HMI tags "Tabla de variables estándar"
   "IndR6" : Bool AT %DB121.DBX3.0, 100 ms
   "IndVparp6" : Bool AT %DB121.DBX70.5, 1 s
   "Auto6" : Bool AT %DB88.DBX10.5, 1 s
   "PanMCH6" : Bool AT %DB88.DBX6.5, 1 s
   "LimSUP6" : Real AT %DB122.DBD20, 1 s
   "LimINF6" : Real AT %DB122.DBD44, 1 s
   "VCMP6" : Int AT %DB125.DBW12, 1 s
   "IncP6" : Bool AT %DB125.DBX16.1, 100 ms
   "DecP6" : Bool AT %DB125.DBX16.7, 1 s
   "SPONF6" : Real AT %DB136.DBD24, 1 s
   "SPOFFF6" : Real AT %DB136.DBD48, 1 s
   "ForzarMarcha6" : Bool AT %DB136.DBX0.5, 1 s
   "ForzarParada6" : Bool AT %DB136.DBX1.3, 1 s
   "ForzandoMarcha6" : Bool AT %DB136.DBX2.1, 1 s
   "SPON6" : Real AT %DB135.DBD32, 1 s
   "SPOFF6" : Real AT %DB135.DBD56, 1 s
   "AnimMenuMC006" : Int AT %DB135.DBW10, 1 s
   "MantMC006" : Bool AT %DB135.DBX60.5, 1 s
   "MarchaOK6" : Bool AT %DB135.DBX61.3, 1 s
   "MarchaMC006" : Bool AT %DB135.DBX62.1, 1 s
   "ParadaMC006" : Bool AT %DB135.DBX62.7, 1 s
   "HORAS6" : DInt AT %DB73.DBD20, 1 s
   "MIN6" : Int AT %DB73.DBW34, 1 s
   "AnimMotorMC006" : Byte AT %DB46.DBB45, 1 s
   "EV6" : Bool AT %Q6.3, 1 s
   "ProxMantMC001_1" : DInt = PLC ProxMantMC001_1 AT %MD768, 1 s
   "ProxMantMC001_2" : DInt = PLC ProxMantMC001_2 AT %MD792, 1 s
   "Varios_UltimoMantMC001_1" : DInt = PLC Varios.UltimoMantMC001_1 AT %DB2.DBD48, 1 s
   "Varios_UltimoMantMC001_2" : DInt = PLC Varios.UltimoMantMC001_2 AT %DB2.DBD72, 1 s
   "ProxMantMC002_1" : DInt = PLC ProxMantMC002_1 AT %MD772, 1 s
   "ProxMantMC002_2" : DInt = PLC ProxMantMC002_2 AT %MD796, 1 s
   "ProxMantMC003_1" : DInt = PLC ProxMantMC003_1 AT %MD776, 1 s
   "ProxMantMC003_2" : DInt = PLC ProxMantMC003_2 AT %MD800, 1 s
   "ProxMantMC004_1" : DInt = PLC ProxMantMC004_1 AT %MD780, 1 s
   "ProxMantMC004_2" : DInt = PLC ProxMantMC004_2 AT %MD804, 1 s
   "ProxMantMC005_1" : DInt = PLC ProxMantMC005_1 AT %MD784, 1 s
   "ProxMantMC005_2" : DInt = PLC ProxMantMC005_2 AT %MD808, 1 s
   "ProxMantMC006_1" : DInt = PLC ProxMantMC006_1 AT %MD788, 1 s
   "ProxMantMC006_2" : DInt = PLC ProxMantMC006_2 AT %MD812, 1 s
   "Varios_UltimoMantMC002_1" : DInt = PLC Varios.UltimoMantMC002_1 AT %DB2.DBD52, 1 s
   "Varios_UltimoMantMC002_2" : DInt = PLC Varios.UltimoMantMC002_2 AT %DB2.DBD76, 1 s
   "Varios_UltimoMantMC003_1" : DInt = PLC Varios.UltimoMantMC003_1 AT %DB2.DBD56, 1 s
   "Varios_UltimoMantMC003_2" : DInt = PLC Varios.UltimoMantMC003_2 AT %DB2.DBD80, 1 s
   "Varios_UltimoMantMC004_1" : DInt = PLC Varios.UltimoMantMC004_1 AT %DB2.DBD60, 1 s
   "Varios_UltimoMantMC004_2" : DInt = PLC Varios.UltimoMantMC004_2 AT %DB2.DBD84, 1 s
   "Varios_UltimoMantMC005_1" : DInt = PLC Varios.UltimoMantMC005_1 AT %DB2.DBD64, 1 s
   "Varios_UltimoMantMC005_2" : DInt = PLC Varios.UltimoMantMC005_2 AT %DB2.DBD88, 1 s
   "Varios_UltimoMantMC006_1" : DInt = PLC Varios.UltimoMantMC006_1 AT %DB2.DBD68, 1 s
   "Varios_UltimoMantMC006_2" : DInt = PLC Varios.UltimoMantMC006_2 AT %DB2.DBD92, 1 s
   "Varios_HorasMantMC001_1" : DInt = PLC Varios.HorasMantMC001_1 AT %DB2.DBD0, 1 s
   "Varios_HorasMantMC006_1" : DInt = PLC Varios.HorasMantMC006_1 AT %DB2.DBD20, 1 s
   "Varios_HorasMantMC006_2" : DInt = PLC Varios.HorasMantMC006_2 AT %DB2.DBD44, 1 s
   "Varios_HorasMantMC002_1" : DInt = PLC Varios.HorasMantMC002_1 AT %DB2.DBD4, 1 s
   "Varios_HorasMantMC001_2" : DInt = PLC Varios.HorasMantMC001_2 AT %DB2.DBD24, 1 s
   "Varios_HorasMantMC002_2" : DInt = PLC Varios.HorasMantMC002_2 AT %DB2.DBD28, 1 s
   "Varios_HorasMantMC004_1" : DInt = PLC Varios.HorasMantMC004_1 AT %DB2.DBD12, 1 s
   "Varios_HorasMantMC004_2" : DInt = PLC Varios.HorasMantMC004_2 AT %DB2.DBD36, 1 s
   "Varios_HorasMantMC005_1" : DInt = PLC Varios.HorasMantMC005_1 AT %DB2.DBD16, 1 s
   "Varios_HorasMantMC005_2" : DInt = PLC Varios.HorasMantMC005_2 AT %DB2.DBD40, 1 s
   "Varios_HorasMantMC003_1" : DInt = PLC Varios.HorasMantMC003_1 AT %DB2.DBD8, 1 s
   "Varios_HorasMantMC003_2" : DInt = PLC Varios.HorasMantMC003_2 AT %DB2.DBD32, 1 s
   "EstadoMantMC003" : Byte = PLC EstadoMantMC003 AT %MB763, 1 s
   "EstadoMantMC005" : Byte = PLC EstadoMantMC005 AT %MB765, 1 s
   "EstadoMantMC004" : Byte = PLC EstadoMantMC004 AT %MB764, 1 s
   "EstadoMantMC002" : Byte = PLC EstadoMantMC002 AT %MB762, 1 s
   "EstadoMantMC001" : Byte = PLC EstadoMantMC001 AT %MB761, 1 s
   "EstadoMantMC006" : Byte = PLC EstadoMantMC006 AT %MB766, 1 s
   "LimiteMantMC001_1" : Bool = PLC LimiteMantMC001_1 AT %M761.0, 1 s
   "LimiteMantMC001_2" : Bool = PLC LimiteMantMC001_2 AT %M761.1, 1 s
   "LimiteMantMC002_1" : Bool = PLC LimiteMantMC002_1 AT %M762.0, 1 s
   "LimiteMantMC002_2" : Bool = PLC LimiteMantMC002_2 AT %M762.1, 1 s
   "LimiteMantMC003_1" : Bool = PLC LimiteMantMC003_1 AT %M763.0, 1 s
   "LimiteMantMC003_2" : Bool = PLC LimiteMantMC003_2 AT %M763.1, 1 s
   "LimiteMantMC004_1" : Bool = PLC LimiteMantMC004_1 AT %M764.0, 1 s
   "LimiteMantMC004_2" : Bool = PLC LimiteMantMC004_2 AT %M764.1, 1 s
   "LimiteMantMC005_1" : Bool = PLC LimiteMantMC005_1 AT %M765.0, 1 s
   "LimiteMantMC005_2" : Bool = PLC LimiteMantMC005_2 AT %M765.1, 1 s
   "LimiteMantMC006_1" : Bool = PLC LimiteMantMC006_1 AT %M766.0, 1 s
   "LimiteMantMC006_2" : Bool = PLC LimiteMantMC006_2 AT %M766.1, 1 s
   "Varios_HorasMantMS050" : DInt = PLC Varios.HorasMantMS050 AT %DB2.DBD96, 1 s
   "Varios_HorasMantMS051" : DInt = PLC Varios.HorasMantMS051 AT %DB2.DBD100, 1 s
   "Varios_HorasMantMS052" : DInt = PLC Varios.HorasMantMS052 AT %DB2.DBD104, 1 s
   "Varios_HorasMantMS053" : DInt = PLC Varios.HorasMantMS053 AT %DB2.DBD108, 1 s
   "HorasSecAlta_HMMS050" : DInt = PLC HorasSecAlta.HMMS050 AT %DB19.DBD0, 1 s
   "HorasSecAlta_HMMS051" : DInt = PLC HorasSecAlta.HMMS051 AT %DB19.DBD4, 1 s
   "HorasSecAlta_HMMS052" : DInt = PLC HorasSecAlta.HMMS052 AT %DB19.DBD8, 1 s
   "HorasSecAlta_HMMS053" : DInt = PLC HorasSecAlta.HMMS053 AT %DB19.DBD12, 1 s
   "Varios_UltimoMantMS050" : DInt = PLC Varios.UltimoMantMS050 AT %DB2.DBD112, 1 s
   "HorasSecAlta_MMMS050" : Int = PLC HorasSecAlta.MMMS050 AT %DB19.DBW16, 1 s
   "ProxMantMS050" : DInt = PLC ProxMantMS050 AT %MD816, 1 s
   "Varios_UltimoMantMS051" : DInt = PLC Varios.UltimoMantMS051 AT %DB2.DBD116, 1 s
   "ProxMantMS051" : DInt = PLC ProxMantMS051 AT %MD820, 1 s
   "HorasSecAlta_MMMS051" : Int = PLC HorasSecAlta.MMMS051 AT %DB19.DBW18, 1 s
   "Varios_UltimoMantMS052" : DInt = PLC Varios.UltimoMantMS052 AT %DB2.DBD120, 1 s
   "ProxMantMS052" : DInt = PLC ProxMantMS052 AT %MD824, 1 s
   "HorasSecAlta_MMMS052" : Int = PLC HorasSecAlta.MMMS052 AT %DB19.DBW20, 1 s
   "Varios_UltimoMantMS053" : DInt = PLC Varios.UltimoMantMS053 AT %DB2.DBD124, 1 s
   "ProxMantMS053" : DInt = PLC ProxMantMS053 AT %MD828, 1 s
   "HorasSecAlta_MMMS053" : Int = PLC HorasSecAlta.MMMS053 AT %DB19.DBW22, 1 s
   "LimiteMantMS051" : Bool = PLC LimiteMantMS051 AT %M767.1, 1 s
   "LimiteMantMS053" : Bool = PLC LimiteMantMS053 AT %M767.3, 1 s
   "LimiteMantMS052" : Bool = PLC LimiteMantMS052 AT %M767.2, 1 s
   "LimiteMantMS050" : Bool = PLC LimiteMantMS050 AT %M767.0, 1 s
   "Varios_HorasMantMC060_1" : DInt = PLC Varios.HorasMantMC060_1 AT %DB2.DBD128, 1 s
   "Varios_HorasMantMC060_2" : DInt = PLC Varios.HorasMantMC060_2 AT %DB2.DBD152, 1 s
   "Varios_HorasMantMC060_3" : DInt = PLC Varios.HorasMantMC060_3 AT %DB2.DBD176, 1 s
   "Varios_HorasMantMC060_4" : DInt = PLC Varios.HorasMantMC060_4 AT %DB2.DBD200, 1 s
   "Varios_UltimoMantMC060_5" : DInt = PLC Varios.UltimoMantMC060_5 AT %DB2.DBD344, 1 s
   "Varios_UltimoMantMC062_1" : DInt = PLC Varios.UltimoMantMC062_1 AT %DB2.DBD256, 1 s
   "Varios_HorasMantMC061_1" : DInt = PLC Varios.HorasMantMC061_1 AT %DB2.DBD132, 1 s
   "Varios_HorasMantMC061_2" : DInt = PLC Varios.HorasMantMC061_2 AT %DB2.DBD156, 1 s
   "Varios_HorasMantMC061_3" : DInt = PLC Varios.HorasMantMC061_3 AT %DB2.DBD180, 1 s
   "Varios_HorasMantMC061_4" : DInt = PLC Varios.HorasMantMC061_4 AT %DB2.DBD204, 1 s
   "Varios_HorasMantMC061_5" : DInt = PLC Varios.HorasMantMC061_5 AT %DB2.DBD228, 1 s
   "Varios_HorasMantMC062_1" : DInt = PLC Varios.HorasMantMC062_1 AT %DB2.DBD136, 1 s
   "Varios_HorasMantMC062_2" : DInt = PLC Varios.HorasMantMC062_2 AT %DB2.DBD160, 1 s
   "Varios_HorasMantMC062_3" : DInt = PLC Varios.HorasMantMC062_3 AT %DB2.DBD184, 1 s
   "Varios_HorasMantMC062_4" : DInt = PLC Varios.HorasMantMC062_4 AT %DB2.DBD208, 1 s
   "Varios_HorasMantMC062_5" : DInt = PLC Varios.HorasMantMC062_5 AT %DB2.DBD232, 1 s
   "Varios_HorasMantMC063_1" : DInt = PLC Varios.HorasMantMC063_1 AT %DB2.DBD140, 1 s
   "Varios_HorasMantMC063_2" : DInt = PLC Varios.HorasMantMC063_2 AT %DB2.DBD164, 1 s
   "Varios_HorasMantMC063_3" : DInt = PLC Varios.HorasMantMC063_3 AT %DB2.DBD188, 1 s
   "Varios_HorasMantMC063_4" : DInt = PLC Varios.HorasMantMC063_4 AT %DB2.DBD212, 1 s
   "Varios_HorasMantMC063_5" : DInt = PLC Varios.HorasMantMC063_5 AT %DB2.DBD236, 1 s
   "Varios_HorasMantMC064_1" : DInt = PLC Varios.HorasMantMC064_1 AT %DB2.DBD144, 1 s
   "Varios_HorasMantMC064_2" : DInt = PLC Varios.HorasMantMC064_2 AT %DB2.DBD168, 1 s
   "Varios_HorasMantMC064_3" : DInt = PLC Varios.HorasMantMC064_3 AT %DB2.DBD192, 1 s
   "Varios_HorasMantMC064_4" : DInt = PLC Varios.HorasMantMC064_4 AT %DB2.DBD216, 1 s
   "Varios_HorasMantMC064_5" : DInt = PLC Varios.HorasMantMC064_5 AT %DB2.DBD240, 1 s
   "Varios_HorasMantMS054_1" : DInt = PLC Varios.HorasMantMS054_1 AT %DB2.DBD368, 1 s
   "Varios_HorasMantMS054_2" : DInt = PLC Varios.HorasMantMS054_2 AT %DB2.DBD380, 1 s
   "Varios_UltimoMantMS055_1" : DInt = PLC Varios.UltimoMantMS055_1 AT %DB2.DBD396, 1 s
   "Varios_HorasMantMS055_2" : DInt = PLC Varios.HorasMantMS055_2 AT %DB2.DBD384, 1 s
   "HorasCmpBaja_HMMC060" : DInt = PLC HorasCmpBaja.HMMC060 AT %DB20.DBD0, 1 s
   "HorasCmpBaja_MMMC060" : Int = PLC HorasCmpBaja.MMMC060 AT %DB20.DBW24, 1 s
   "Varios_UltimoMantMC060_1" : DInt = PLC Varios.UltimoMantMC060_1 AT %DB2.DBD248, 1 s
   "ProxMantMC060_1" : DInt = PLC ProxMantMC060_1 AT %MD834, 1 s
   "ProxMantMC060_2" : DInt = PLC ProxMantMC060_2 AT %MD858, 1 s
   "ProxMantMC060_3" : DInt = PLC ProxMantMC060_3 AT %MD882, 1 s
   "ProxMantMC060_4" : DInt = PLC ProxMantMC060_4 AT %MD918, 1 s
   "ProxMantMC060_5" : DInt = PLC ProxMantMC060_5 AT %MD942, 1 s
   "Varios_UltimoMantMC060_2" : DInt = PLC Varios.UltimoMantMC060_2 AT %DB2.DBD272, 1 s
   "Varios_UltimoMantMC060_3" : DInt = PLC Varios.UltimoMantMC060_3 AT %DB2.DBD296, 1 s
   "Varios_UltimoMantMC060_4" : DInt = PLC Varios.UltimoMantMC060_4 AT %DB2.DBD320, 1 s
   "HorasCmpBaja_HMMC061" : DInt = PLC HorasCmpBaja.HMMC061 AT %DB20.DBD4, 1 s
   "ProxMantMC061_1" : DInt = PLC ProxMantMC061_1 AT %MD838, 1 s
   "ProxMantMC061_3" : DInt = PLC ProxMantMC061_3 AT %MD886, 1 s
   "ProxMantMC061_4" : DInt = PLC ProxMantMC061_4 AT %MD922, 1 s
   "ProxMantMC061_2" : DInt = PLC ProxMantMC061_2 AT %MD862, 1 s
   "ProxMantMC061_5" : DInt = PLC ProxMantMC061_5 AT %MD946, 1 s
   "Varios_UltimoMantMC061_1" : DInt = PLC Varios.UltimoMantMC061_1 AT %DB2.DBD252, 1 s
   "Varios_UltimoMantMC061_2" : DInt = PLC Varios.UltimoMantMC061_2 AT %DB2.DBD276, 1 s
   "Varios_UltimoMantMC061_3" : DInt = PLC Varios.UltimoMantMC061_3 AT %DB2.DBD300, 1 s
   "Varios_UltimoMantMC061_4" : DInt = PLC Varios.UltimoMantMC061_4 AT %DB2.DBD324, 1 s
   "Varios_UltimoMantMC061_5" : DInt = PLC Varios.UltimoMantMC061_5 AT %DB2.DBD348, 1 s
   "HorasCmpBaja_MMMC061" : Int = PLC HorasCmpBaja.MMMC061 AT %DB20.DBW26, 1 s
   "HorasCmpBaja_HMMC062" : DInt = PLC HorasCmpBaja.HMMC062 AT %DB20.DBD8, 1 s
   "HorasCmpBaja_MMMC062" : Int = PLC HorasCmpBaja.MMMC062 AT %DB20.DBW28, 1 s
   "ProxMantMC062_1" : DInt = PLC ProxMantMC062_1 AT %MD842, 1 s
   "ProxMantMC062_2" : DInt = PLC ProxMantMC062_2 AT %MD866, 1 s
   "ProxMantMC062_3" : DInt = PLC ProxMantMC062_3 AT %MD890, 1 s
   "ProxMantMC062_4" : DInt = PLC ProxMantMC062_4 AT %MD926, 1 s
   "ProxMantMC062_5" : DInt = PLC ProxMantMC062_5 AT %MD950, 1 s
   "Varios_UltimoMantMC062_5" : DInt = PLC Varios.UltimoMantMC062_5 AT %DB2.DBD352, 1 s
   "Varios_UltimoMantMC062_3" : DInt = PLC Varios.UltimoMantMC062_3 AT %DB2.DBD304, 1 s
   "Varios_UltimoMantMC062_2" : DInt = PLC Varios.UltimoMantMC062_2 AT %DB2.DBD280, 1 s
   "HorasCmpBaja_HMMC063" : DInt = PLC HorasCmpBaja.HMMC063 AT %DB20.DBD12, 1 s
   "HorasCmpBaja_MMMC063" : Int = PLC HorasCmpBaja.MMMC063 AT %DB20.DBW30, 1 s
   "ProxMantMC063_1" : DInt = PLC ProxMantMC063_1 AT %MD846, 1 s
   "ProxMantMC063_2" : DInt = PLC ProxMantMC063_2 AT %MD870, 1 s
   "ProxMantMC063_3" : DInt = PLC ProxMantMC063_3 AT %MD894, 1 s
   "ProxMantMC063_4" : DInt = PLC ProxMantMC063_4 AT %MD930, 1 s
   "ProxMantMC063_5" : DInt = PLC ProxMantMC063_5 AT %MD954, 1 s
   "HorasCmpBaja_HMMC064" : DInt = PLC HorasCmpBaja.HMMC064 AT %DB20.DBD16, 1 s
   "Varios_UltimoMantMC063_1" : DInt = PLC Varios.UltimoMantMC063_1 AT %DB2.DBD260, 1 s
   "Varios_UltimoMantMC063_2" : DInt = PLC Varios.UltimoMantMC063_2 AT %DB2.DBD284, 1 s
   "Varios_UltimoMantMC063_3" : DInt = PLC Varios.UltimoMantMC063_3 AT %DB2.DBD308, 1 s
   "Varios_UltimoMantMC063_4" : DInt = PLC Varios.UltimoMantMC063_4 AT %DB2.DBD332, 1 s
   "Varios_UltimoMantMC063_5" : DInt = PLC Varios.UltimoMantMC063_5 AT %DB2.DBD356, 1 s
   "HorasCmpBaja_MMMC064" : Int = PLC HorasCmpBaja.MMMC064 AT %DB20.DBW32, 1 s
   "ProxMantMC064_1" : DInt = PLC ProxMantMC064_1 AT %MD850, 1 s
   "ProxMantMC064_2" : DInt = PLC ProxMantMC064_2 AT %MD874, 1 s
   "ProxMantMC064_3" : DInt = PLC ProxMantMC064_3 AT %MD910, 1 s
   "ProxMantMC064_4" : DInt = PLC ProxMantMC064_4 AT %MD934, 1 s
   "ProxMantMC064_5" : DInt = PLC ProxMantMC064_5 AT %MD958, 1 s
   "Varios_UltimoMantMC064_1" : DInt = PLC Varios.UltimoMantMC064_1 AT %DB2.DBD264, 1 s
   "Varios_UltimoMantMC064_5" : DInt = PLC Varios.UltimoMantMC064_5 AT %DB2.DBD360, 1 s
   "Varios_UltimoMantMC064_2" : DInt = PLC Varios.UltimoMantMC064_2 AT %DB2.DBD288, 1 s
   "Varios_UltimoMantMC064_3" : DInt = PLC Varios.UltimoMantMC064_3 AT %DB2.DBD312, 1 s
   "Varios_UltimoMantMC064_4" : DInt = PLC Varios.UltimoMantMC064_4 AT %DB2.DBD336, 1 s
   "LimiteMantMC060_1" : Bool = PLC LimiteMantMC060_1 AT %M901.0, 1 s
   "LimiteMantMC060_2" : Bool = PLC LimiteMantMC060_2 AT %M901.1, 1 s
   "LimiteMantMC060_3" : Bool = PLC LimiteMantMC060_3 AT %M901.2, 1 s
   "LimiteMantMC060_4" : Bool = PLC LimiteMantMC060_4 AT %M901.3, 1 s
   "LimiteMantMC060_5" : Bool = PLC LimiteMantMC060_5 AT %M901.4, 1 s
   "EstadoMantMC060" : Byte = PLC EstadoMantMC060 AT %MB901, 1 s
   "EstadoMantMC061" : Byte = PLC EstadoMantMC061 AT %MB902, 1 s
   "EstadoMantMC062" : Byte = PLC EstadoMantMC062 AT %MB903, 1 s
   "EstadoMantMC063" : Byte = PLC EstadoMantMC063 AT %MB904, 1 s
   "EstadoMantMC064" : Byte = PLC EstadoMantMC064 AT %MB905, 1 s
   "HorasSecBaja_HMMS054" : DInt = PLC HorasSecBaja.HMMS054 AT %DB24.DBD0, 1 s
   "HorasSecBaja_MMMS054" : Int = PLC HorasSecBaja.MMMS054 AT %DB24.DBW12, 1 s
   "ProxMantMS054_1" : DInt = PLC ProxMantMS054_1 AT %MD966, 1 s
   "ProxMantMS054_2" : DInt = PLC ProxMantMS054_2 AT %MD970, 1 s
   "Varios_UltimoMantMS054_1" : DInt = PLC Varios.UltimoMantMS054_1 AT %DB2.DBD392, 1 s
   "Varios_UltimoMantMS054_2" : DInt = PLC Varios.UltimoMantMS054_2 AT %DB2.DBD404, 1 s
   "EstadoMantSecBaja" : Byte = PLC EstadoMantSecBaja AT %MB832, 1 s
   "LimiteMantMS054_1" : Bool = PLC LimiteMantMS054_1 AT %M832.0, 1 s
   "LimiteMantMS054_2" : Bool = PLC LimiteMantMS054_2 AT %M832.1, 1 s
   "LimiteMantMS055_1" : Bool = PLC LimiteMantMS055_1 AT %M832.2, 1 s
   "LimiteMantMS055_2" : Bool = PLC LimiteMantMS055_2 AT %M832.3, 1 s
   "HorasSecBaja_HMMS055" : DInt = PLC HorasSecBaja.HMMS055 AT %DB24.DBD4, 1 s
   "HorasSecBaja_MMMS055" : Int = PLC HorasSecBaja.MMMS055 AT %DB24.DBW14, 1 s
   "ProxMantMS055_1" : DInt = PLC ProxMantMS055_1 AT %MD974, 1 s
   "ProxMantMS055_2" : DInt = PLC ProxMantMS055_2 AT %MD978, 1 s
   "Varios_UltimoMantMS055_2" : DInt = PLC Varios.UltimoMantMS055_2 AT %DB2.DBD408, 1 s
   "Varios_HorasMantBost1" : DInt = PLC Varios.HorasMantBost1 AT %DB2.DBD416, 1 s
   "Varios_HorasMantBost2" : DInt = PLC Varios.HorasMantBost2 AT %DB2.DBD420, 1 s
   "ProxMantBoost1" : DInt = PLC ProxMantBoost1 AT %MD16, 1 s
   "ProxMantBoost2" : DInt = PLC ProxMantBoost2 AT %MD26, 1 s
   "Varios_UltimoMantBoost1" : DInt = PLC Varios.UltimoMantBoost1 AT %DB2.DBD424, 1 s
   "Varios_UltimoMantBoost2" : DInt = PLC Varios.UltimoMantBoost2 AT %DB2.DBD428, 1 s
   "LimiteMantBoost1" : Bool = PLC LimiteMantBoost1 AT %M1.7, 1 s
   "LimiteMantBoost2" : Bool = PLC LimiteMantBoost2 AT %M2.3, 1 s
   "DBParamCmpALTA-MTA_TempCritEnclav" : Real = PLC "DBParamCmpALTA-MTA".TempCritEnclav AT %DB122.DBD100, 1 s
   "NumeroCompresor" : Int, internal
   "EstadoRegistro" : Bool, internal
   "DB-PurgaComAlta_Habil_PurgaBallis" : Bool = PLC "DB-PurgaComAlta".Habil_PurgaBellis AT %DB53.DBX0.0, 1 s
   "DB-PurgaComAlta_Toff_PurgaBallis" : Word = PLC "DB-PurgaComAlta".Toff_PurgaBellis AT %DB53.DBW2, 1 s
   "DB-PurgaComAlta_Ton_PurgaBallis" : Word = PLC "DB-PurgaComAlta".Ton_PurgaBellis AT %DB53.DBW4, 1 s
   "DB-PurgaComAlta_Habil_PurgaABC2" : Bool = PLC "DB-PurgaComAlta".Habil_PurgaABC2 AT %DB53.DBX0.1, 1 s
   "DB-PurgaComAlta_Toff_PurgaABC2" : Word = PLC "DB-PurgaComAlta".Toff_PurgaABC2 AT %DB53.DBW6, 1 s
   "DB-PurgaComAlta_Ton_PurgaABC2" : Word = PLC "DB-PurgaComAlta".Ton_PurgaABC2 AT %DB53.DBW8, 1 s
   "DB-PurgaComAlta_Habil_PurgaABC3" : Bool = PLC "DB-PurgaComAlta".Habil_PurgaABC3 AT %DB53.DBX0.2, 1 s
   "DB-PurgaComAlta_Toff_PurgaABC3" : Word = PLC "DB-PurgaComAlta".Toff_PurgaABC3 AT %DB53.DBW10, 1 s
   "DB-PurgaComAlta_Ton_PurgaABC3" : Word = PLC "DB-PurgaComAlta".Ton_PurgaABC3 AT %DB53.DBW12, 1 s
   "DB-PurgaComAlta_Habil_PurgaABC4" : Bool = PLC "DB-PurgaComAlta".Habil_PurgaABC4 AT %DB53.DBX0.3, 1 s
   "DB-PurgaComAlta_Toff_PurgaABC4" : Word = PLC "DB-PurgaComAlta".Toff_PurgaABC4 AT %DB53.DBW14, 1 s
   "DB-PurgaComAlta_Ton_PurgaABC4" : Word = PLC "DB-PurgaComAlta".Ton_PurgaABC4 AT %DB53.DBW16, 1 s
   "DB-PurgaComAlta_Habil_PurgaABC5" : Bool = PLC "DB-PurgaComAlta".Habil_PurgaABC5 AT %DB53.DBX0.4, 1 s
   "DB-PurgaComAlta_Toff_PurgaABC5" : Word = PLC "DB-PurgaComAlta".Toff_PurgaABC5 AT %DB53.DBW18, 1 s
   "DB-PurgaComAlta_Ton_PurgaABC5" : Word = PLC "DB-PurgaComAlta".Ton_PurgaABC5 AT %DB53.DBW20, 1 s
   "DB-PurgaComAlta_Habil_PurgaABC1" : Bool = PLC "DB-PurgaComAlta".Habil_PurgaABC1 AT %DB53.DBX0.5, 1 s
   "DB-PurgaComAlta_Toff_PurgaABC1" : Word = PLC "DB-PurgaComAlta".Toff_PurgaABC1 AT %DB53.DBW22, 1 s
   "DB-PurgaComAlta_Ton_PurgaABC1" : Word = PLC "DB-PurgaComAlta".Ton_PurgaABC1 AT %DB53.DBW24, 1 s
   "DB-PurgaComAlta_Prueba_PurgaBallis" : Bool = PLC "DB-PurgaComAlta".Prueba_PurgaBellis AT %DB53.DBX26.0, 1 s
   "MC003_EVP" : Bool = PLC MC003_EVP AT %Q7.2, 1 s
   "MC001_EVP" : Bool = PLC MC001_EVP AT %Q7.3, 1 s
   "MC002_EVP" : Bool = PLC MC002_EVP AT %Q7.4, 1 s
   "MC004_EVP" : Bool = PLC MC004_EVP AT %Q7.5, 1 s
   "MC005_EVP" : Bool = PLC MC005_EVP AT %Q7.6, 1 s
   "MC006_EVP" : Bool = PLC MC006_EVP AT %Q7.7, 1 s
   "DB-PurgaComAlta_Prueba_PurgaABC2" : Bool = PLC "DB-PurgaComAlta".Prueba_PurgaABC2 AT %DB53.DBX26.1, 1 s
   "DB-PurgaComAlta_Prueba_PurgaABC3" : Bool = PLC "DB-PurgaComAlta".Prueba_PurgaABC3 AT %DB53.DBX26.2, 1 s
   "DB-PurgaComAlta_Prueba_PurgaABC4" : Bool = PLC "DB-PurgaComAlta".Prueba_PurgaABC4 AT %DB53.DBX26.3, 1 s
   "DB-PurgaComAlta_Prueba_PurgaABC5" : Bool = PLC "DB-PurgaComAlta".Prueba_PurgaABC5 AT %DB53.DBX26.4, 1 s
   "DB-PurgaComAlta_Prueba_PurgaABC1" : Bool = PLC "DB-PurgaComAlta".Prueba_PurgaABC1 AT %DB53.DBX26.5, 1 s
   "DB_ALA_MEM_x199" : Bool = PLC DB_ALA_MEM.x199 AT %DB34.DBX24.7, 1 s
   "Enclavamientos_En1" : Bool = PLC Enclavamientos.En1 AT %DB28.DBX0.0, 1 s   // Encl de compresores por flujostato
   "Enclavamientos_En2" : Bool = PLC Enclavamientos.En2 AT %DB28.DBX0.1, 1 s   // Encl de compresores por temperatura

HMI tags "Tabla de variables estándar_1"
   "MC066_STD" : Real AT %DB14.DBD26, 1 s
   "MV031_STD" : Word AT %DB14.DBW70, 1 s
   "MV032_STD" : Word AT %DB14.DBW72, 1 s
   "MV030_STD" : Word AT %DB14.DBW68, 1 s
   "DIP_1" : Int, internal
   "MP016_STD" : Word AT %DB14.DBW40, 1 s
   "MC004_STD" : Word AT %DB14.DBW8, 1 s
   "MP013_STD" : Word AT %DB14.DBW34, 1 s
   "MV033_STD" : Word AT %DB14.DBW74, 1 s
   "MC001_STD" : Word AT %DB14.DBW2, 1 s
   "MC060_STD" : Word AT %DB14.DBW14, 1 s
   "MC002_STD" : Word AT %DB14.DBW4, 1 s
   "MP012_STD" : Word AT %DB14.DBW32, 1 s
   "MC065_STD" : Word AT %DB14.DBW24, 1 s
   "MS051_STD" : Word AT %DB14.DBW50, 1 s
   "MC006_STD" : Word AT %DB14.DBW12, 1 s
   "MP011_STD" : Word AT %DB14.DBW30, 1 s
   "Iluminati_STD" : Word AT %DB14.DBW60, 1 s
   "MC064_STD" : Word AT %DB14.DBW22, 1 s
   "MS052_STD" : Word AT %DB14.DBW52, 1 s
   "MT010_STD" : Word AT %DB14.DBW42, 1 s
   "MS053_STD" : Word AT %DB14.DBW54, 1 s
   "MP019_STD" : Word AT %DB14.DBW46, 1 s
   "MC005_STD" : Word AT %DB14.DBW10, 1 s
   "MC061_STD" : Word AT %DB14.DBW16, 1 s
   "MV034_STD" : Word AT %DB14.DBW76, 1 s
   "MC063_STD" : Word AT %DB14.DBW20, 1 s
   "MP015_STD" : Word AT %DB14.DBW38, 1 s
   "MT007_STD" : Word AT %DB14.DBW62, 1 s
   "MS055_STD" : Word AT %DB14.DBW58, 1 s
   "MP018_STD" : Word AT %DB14.DBW44, 1 s
   "MP014_STD" : Word AT %DB14.DBW36, 1 s
   "MS054_STD" : Word AT %DB14.DBW56, 1 s
   "MS050_STD" : Word AT %DB14.DBW48, 1 s
   "MP010_STD" : Word AT %DB14.DBW28, 1 s
   "MT008_STD" : Word AT %DB14.DBW64, 1 s
   "MT009_STD" : Word AT %DB14.DBW66, 1 s
   "MC003_STD" : Word AT %DB14.DBW6, 1 s
   "MC062_STD" : Word AT %DB14.DBW18, 1 s
   "EB5" : Word AT %MW5, 1 s
   "EB7" : Word AT %MW7, 1 s
   "EB4" : Word AT %MW4, 1 s
   "EW8" : Word AT %MW22, 1 s
   "ACK_ALARMA_2" : Int AT %DB40.DBW0, 1 s
   "MP020_STD" : Word AT %DB14.DBW78, 1 s
   "MP021_STD" : Word AT %DB14.DBW80, 1 s
   "MP022_STD" : Word AT %DB14.DBW82, 1 s
   "CERO" : Bool AT %M0.0, 1 s
   "UNO" : Bool AT %M0.1, 1 s
   "IndCh" : Bool AT %M310.0, 1 s
   "IndTrCh" : Bool AT %M310.1, 1 s
   "IndCmpBaja" : Bool AT %M310.2, 1 s
   "IndSecBaja" : Bool AT %M310.3, 1 s
   "IndCmpAlta" : Bool AT %M310.4, 1 s
   "IndSecAlta" : Bool AT %M310.5, 1 s
   "IndTrCav" : Bool AT %M310.6, 1 s
   "AnularSirena?" : Bool, internal
   "HorasBoost1" : DInt AT %DB62.DBD8, 1 s
   "HorasBoost2" : DInt AT %DB62.DBD12, 1 s
   "BoostPrHoras" : Bool AT %M330.2, 1 s
   "BoostInvP" : Bool AT %M330.1, 1 s
   "PrioridadBoost1" : Int AT %MW332, 1 s
   "PrioridadBoost2" : Int AT %MW334, 1 s
   "BoostInvPMan" : Bool AT %M330.3, 1 s
   "min_boost1" : Int AT %DB62.DBW4, 1 s
   "SegsBoost1" : Int AT %DB62.DBW0, 1 s
   "SegsBoost" : Int AT %DB62.DBW2, 1 s
   "MinBoost2" : Int AT %DB62.DBW6, 1 s
   "FT1_AGUA" : Bool = PLC FT1_AGUA AT %I8.0, 1 s

HMI tags "AlarmasMTA"
   "AlarmasWord0" : Int AT %DB86.DBW0, 1 s
   "AlarmasWord1" : Int AT %DB86.DBW2, 1 s
   "AlarmasWord2" : Int AT %DB86.DBW4, 1 s
   "AlarmasWord3" : Int AT %DB86.DBW6, 1 s
   "AlarmasWord4" : Int AT %DB86.DBW8, 1 s
   "AlarmasWord5" : Int AT %DB86.DBW10, 1 s
   "AlarmasWord6" : Int AT %DB86.DBW12, 1 s
   "AlarmasWord7" : Int AT %DB86.DBW14, 1 s
   "AlarmasWord8" : Int AT %DB86.DBW16, 1 s
   "Rec0" : Int AT %DB86.DBW0, 1 s
   "Rec1" : Int AT %DB86.DBW2, 1 s
   "Rec2" : Int AT %DB86.DBW4, 1 s
   "Rec3" : Int AT %DB86.DBW6, 1 s
   "Rec4" : Int AT %DB86.DBW8, 1 s
   "Rec5" : Int AT %DB86.DBW10, 1 s
   "Rec6" : Int AT %DB86.DBW12, 1 s
   "Rec7" : Int AT %DB86.DBW14, 1 s
   "Rec8" : Int AT %DB86.DBW16, 1 s
   "AlarmasWord9" : Int AT %DB86.DBW18, 1 s
   "AlarmasWord10" : Int AT %DB86.DBW20, 1 s
   "AlarmasWord11" : Int AT %DB86.DBW22, 1 s
   "AlarmasWord12" : Int AT %DB86.DBW24, 1 s
   "AlarmasWord13" : Int AT %DB86.DBW26, 1 s
   "AlarmasWord14" : Int AT %DB86.DBW28, 1 s
   "Rec9" : Int AT %DB86.DBW18, 1 s
   "Rec10" : Int AT %DB86.DBW20, 1 s
   "Rec11" : Int AT %DB86.DBW22, 1 s
   "Rec12" : Int AT %DB86.DBW24, 1 s
   "Rec13" : Int AT %DB86.DBW26, 1 s
   "Rec14" : Int AT %DB86.DBW28, 1 s
   "AlarmasWord15" : Int AT %DB86.DBW30, 1 s
   "Rec15" : Int AT %DB86.DBW30, 1 s
   "ReconocerTODAS" : Bool AT %DB47.DBX0.7, 1 s
   "EncendidoPLC" : Bool AT %M300.1, 1 s
      on ChangeValue: ActivateScreen("INICIO", 0)
   "AlarmasWord16" : Int AT %DB86.DBW32, 1 s
   "Rec16" : Int AT %DB86.DBW32, 1 s
   "ReconocerTODAS_1" : Bool AT %DB47.DBX1.0, 1 s
   "AlarmasWord18" : Int AT %DB86.DBW36, 1 s
   "Rec18" : Int AT %DB86.DBW36, 1 s
   "AlarmasWord19" : Int AT %DB86.DBW38, 1 s
   "Rec19" : Int AT %DB86.DBW38, 1 s
   "AlarmasWord20" : Int AT %DB86.DBW40, 1 s
   "AlarmasWord21" : Int AT %DB86.DBW42, 1 s
   "AlarmasWord22" : Int AT %DB86.DBW44, 1 s
   "AlarmasWord23" : Int AT %DB86.DBW46, 1 s
   "AlarmasWord24" : Int AT %DB86.DBW48, 1 s
   "Rec20" : Int AT %DB86.DBW40, 1 s
   "Rec21" : Int AT %DB86.DBW42, 1 s
   "Rec22" : Int AT %DB86.DBW44, 1 s
   "Rec23" : Int AT %DB86.DBW46, 1 s
   "Rec24" : Int AT %DB86.DBW48, 1 s
   "AlarmasWord17" : Int AT %DB86.DBW34, 1 s
   "Rec17" : Int AT %DB86.DBW34, 1 s

HMI tags "AutoTorresCav"
   "AutoV030" : Bool AT %DB21.DBX6.4, 1 s
   "AutoV031" : Bool AT %DB21.DBX6.5, 1 s
   "SP-OFF-V030" : Int AT %DB21.DBW12, 1 s
   "SP-OFF-V031" : Int AT %DB21.DBW14, 1 s
   "SP-ON-V030" : Int AT %DB21.DBW8, 1 s
   "SP-ON-V031" : Int AT %DB21.DBW10, 1 s

HMI tags "AutoTorresChillers"
   "AutoV001" : Bool AT %DB92.DBX0.0, 1 s
   "AutoV002" : Bool AT %DB92.DBX0.1, 1 s
   "AutoV003" : Bool AT %DB92.DBX0.2, 1 s
   "SP-ON-V001" : Int AT %DB92.DBW2, 1 s
   "SP-ON-V002" : Int AT %DB92.DBW4, 1 s
   "SP-ON-V003" : Int AT %DB92.DBW6, 1 s
   "SP-OFF-V001" : Int AT %DB92.DBW8, 1 s
   "SP-OFF-V002" : Int AT %DB92.DBW10, 1 s
   "SP-OFF-V003" : Int AT %DB92.DBW12, 1 s
   "TemperaturatorresCH" : Real AT %DB52.DBD4, 1 s

HMI tags "Booster"
   "AlarmaBooster" : Bool AT %M10.3, 1 s
   "Booster_ModoManten" : Bool AT %M10.0, 1 s
   "Booster_ModoManual" : Bool AT %M10.1, 1 s
   "Booster_ModoAutoma" : Bool AT %M10.2, 1 s
   "Booster_PlsManten" : Bool AT %M10.5, 1 s
   "Booster_PlsManual" : Bool AT %M10.6, 1 s
   "Booster_PlsAutoma" : Bool AT %M10.7, 1 s
   "AnimaMotBooster" : Byte AT %MB11, 1 s
   "BoosterOrdMarcha" : Bool AT %M10.4, 1 s
   "Booster_Conf_Marcha" : Bool AT %E3.7, 1 s
   "Booster_Presost_Ctrl" : Bool AT %E7.6, 1 s
   "Booster_Presost_PA" : Bool AT %E7.7, 1 s
   "Booster_Habilitacion" : Bool AT %M12.0, 1 s
   "Booster2_Conf_Marcha" : Bool AT %I9.6, 1 s
   "Booster2_Habilitacion" : Bool AT %M13.1, 1 s
   "Booster2_ModoAutoma" : Bool AT %M12.3, 1 s
   "Booster2_ModoManten" : Bool AT %M12.1, 1 s
   "Booster2_ModoManual" : Bool AT %M12.2, 1 s
   "Booster2_PlsAutoma" : Bool AT %M13.0, 1 s
   "Booster2_PlsManten" : Bool AT %M12.6, 1 s
   "Booster2_PlsManual" : Bool AT %M12.7, 1 s
   "AnimaMotBooster2" : Byte AT %MB14, 1 s
   "Booster2OrdMarcha" : Bool AT %M12.5, 1 s
   "TiempoAyudaON" : Int AT %DB62.DBW20, 1 s
   "TiempoAyudaOFF" : Int AT %DB62.DBW22, 1 s
   "DifHorINVBoost" : DInt AT %DB62.DBD16, 1 s
   "LimArrBoostPrio2" : Real AT %DB62.DBD28, 1 s
   "LimArrBoostPrio1" : Real AT %DB62.DBD32, 1 s
   "LimParBoostPrio2" : Real AT %DB62.DBD36, 1 s
   "LimParBoostPrio1" : Real AT %DB62.DBD40, 1 s
   "Presión_Actual_Boosters" : Real AT %MD56, 1 s
   "Ctrl_Analógico" : Bool AT %DB62.DBX44.0, 1 s
   "Ver_Config" : Bool, internal
   "CotaSupPresAna" : Real AT %MD76, 1 s

HMI tags "CFG-Analog-MTA"
   "PresiónALTA" : Real AT %DB52.DBD52, 1 s
   "PresiónBAJA" : Real AT %DB52.DBD16, 1 s
   "TempCAV" : Real AT %DB52.DBD0, 1 s
   "TempCH" : Real AT %DB52.DBD4, 1 s
   "CFG-ALtaHH" : Real AT %DB52.DBD20, 1 s
   "CFG-ALtaH" : Real AT %DB52.DBD24, 1 s
   "CFG-ALtaL" : Real AT %DB52.DBD28, 1 s
   "CFG-ALtaLL" : Real AT %DB52.DBD32, 1 s
   "CFG-BajaHH" : Real AT %DB52.DBD36, 1 s
   "CFG-BajaH" : Real AT %DB52.DBD40, 1 s
   "CFG-BajaL" : Real AT %DB52.DBD44, 1 s
   "CFG-BajaLL" : Real AT %DB52.DBD48, 1 s
   "LO_potencia" : Real = PLC CaudalPotencia.LO_potencia AT %DB26.DBD20, 1 s
   "HI_caudal" : Real = PLC CaudalPotencia.HI_caudal AT %DB26.DBD8, 1 s
   "LO_caudal" : Real = PLC CaudalPotencia.LO_caudal AT %DB26.DBD12, 1 s
   "HI_potencia" : Real = PLC CaudalPotencia.HI_potencia AT %DB26.DBD16, 1 s
   "Caudal" : Real = PLC CaudalPotencia.lecCaudal AT %DB26.DBD0, 1 s
   "Potencia" : Real = PLC CaudalPotencia.lecPotencia AT %DB26.DBD4, 1 s

HMI tags "ChillersMTA"
   "HabMT007" : Bool AT %DB90.DBX6.4, 1 s
   "HabMT008" : Bool AT %DB90.DBX6.5, 1 s
   "HabMT009" : Bool AT %DB90.DBX6.6, 1 s
   "HabMT010" : Bool AT %DB90.DBX6.7, 1 s
   "DesMT007" : Bool AT %DB90.DBX8.1, 1 s
   "DesMT008" : Bool AT %DB90.DBX8.2, 1 s
   "DesMT009" : Bool AT %DB90.DBX8.3, 1 s
   "DesMT010" : Bool AT %DB90.DBX8.4, 1 s
   "MarchaMT007" : Bool AT %DB90.DBX9.6, 1 s
   "MarchaMT008" : Bool AT %DB90.DBX9.7, 1 s
   "MarchaMT009" : Bool AT %DB90.DBX10.0, 1 s
   "MarchaMT010" : Bool AT %DB90.DBX10.1, 1 s
   "ParadaMT007" : Bool AT %DB90.DBX11.3, 1 s
   "ParadaMT008" : Bool AT %DB90.DBX11.4, 1 s
   "ParadaMT009" : Bool AT %DB90.DBX11.5, 1 s
   "ParadaMT010" : Bool AT %DB90.DBX11.6, 1 s
   "Habilitación-CH-SOP-GR" : Bool AT %Q69.4, 1 s
   "Habilitación-CH-SOP-CH" : Bool AT %Q69.5, 1 s
   "Habilitación-CH-ENV-GR" : Bool AT %Q69.6, 1 s
   "Habilitación-CH-ENV-CH" : Bool AT %Q69.7, 1 s
   "Alarma1-CH-SOP-GR" : Bool AT %I68.4, 1 s
   "Alarma2-CH-SOP-GR" : Bool AT %I68.5, 1 s
   "RUN-CH-SOP-GR" : Bool AT %I68.6, 1 s
   "MAX-CH-SOP-GR" : Bool AT %I68.7, 1 s
   "AnimaciónMT007" : Byte AT %DB46.DBB6, 1 s
   "AnimaciónMT008" : Byte AT %DB46.DBB7, 1 s
   "AnimaciónMT009" : Byte AT %DB46.DBB8, 1 s
   "AnimaciónMT010" : Byte AT %DB46.DBB9, 1 s
   "AnimaciónMP010" : Byte AT %DB46.DBB0, 1 s
   "AnimaciónMP011" : Byte AT %DB46.DBB1, 1 s
   "AnimaciónMP012" : Byte AT %DB46.DBB2, 1 s
   "AnimaciónMP013" : Byte AT %DB46.DBB3, 1 s
   "HabMP010" : Bool AT %DB90.DBX7.0, 1 s
   "HabMP011" : Bool AT %DB90.DBX7.1, 1 s
   "HabMP012" : Bool AT %DB90.DBX7.2, 1 s
   "HabMP013" : Bool AT %DB90.DBX7.3, 1 s
   "HabMP018" : Bool AT %DB90.DBX7.4, 1 s
   "HabMP019" : Bool AT %DB90.DBX7.5, 1 s
   "DesMP010" : Bool AT %DB90.DBX8.5, 1 s
   "DesMP011" : Bool AT %DB90.DBX8.6, 1 s
   "DesMP012" : Bool AT %DB90.DBX8.7, 1 s
   "DesMP013" : Bool AT %DB90.DBX9.0, 1 s
   "DesMP018" : Bool AT %DB90.DBX9.1, 1 s
   "DesMP019" : Bool AT %DB90.DBX9.2, 1 s
   "MarchaMP010" : Bool AT %DB90.DBX10.2, 1 s
   "MarchaMP011" : Bool AT %DB90.DBX10.3, 1 s
   "MarchaMP012" : Bool AT %DB90.DBX10.4, 1 s
   "MarchaMP013" : Bool AT %DB90.DBX10.5, 1 s
   "MarchaMP018" : Bool AT %DB90.DBX10.6, 1 s
   "MarchaMP019" : Bool AT %DB90.DBX10.7, 1 s
   "ParadaMP010" : Bool AT %DB90.DBX11.7, 1 s
   "ParadaMP011" : Bool AT %DB90.DBX12.0, 1 s
   "ParadaMP012" : Bool AT %DB90.DBX12.1, 1 s
   "ParadaMP013" : Bool AT %DB90.DBX12.2, 1 s
   "ParadaMP018" : Bool AT %DB90.DBX12.3, 1 s
   "ParadaMP019" : Bool AT %DB90.DBX12.4, 1 s
   "AnimaciónMP018" : Byte AT %DB46.DBB4, 1 s
   "AnimaciónMP019" : Byte AT %DB46.DBB5, 1 s
   "DesV001" : Bool AT %DB90.DBX9.3, 1 s
   "DesV002" : Bool AT %DB90.DBX9.4, 1 s
   "HabV001" : Bool AT %DB90.DBX7.6, 1 s
   "HabV002" : Bool AT %DB90.DBX7.7, 1 s
   "MarchaV001" : Bool AT %DB90.DBX11.0, 1 s
   "MarchaV002" : Bool AT %DB90.DBX11.1, 1 s
   "ParadaV001" : Bool AT %DB90.DBX12.5, 1 s
   "ParadaV002" : Bool AT %DB90.DBX12.6, 1 s
   "AnimaciónV001" : Byte AT %DB46.DBB10, 1 s
   "AnimaciónV002" : Byte AT %DB46.DBB11, 1 s
   "VentiladoresMTA" : Bool, internal
   "MAX-CH-ENV-GR" : Bool AT %I69.7, 1 s
   "RUN-CH-ENV-GR" : Bool AT %I69.6, 1 s
   "Alarma2-CH-ENV-GR" : Bool AT %I69.5, 1 s
   "Alarma1-CH-ENV-GR" : Bool AT %I69.4, 1 s
   "SirenaM1" : Bool AT %DB91.DBX0.0, 1 s
   "SirenaM2" : Bool AT %DB91.DBX0.1, 1 s
   "SirenaM3" : Bool AT %DB91.DBX0.2, 1 s
   "SirenaM4" : Bool AT %DB91.DBX0.3, 1 s
   "AnimaciónV003" : Byte AT %DB46.DBB12, 1 s
   "HabV003" : Bool AT %DB90.DBX8.0, 1 s
   "DesV003" : Bool AT %DB90.DBX9.5, 1 s
   "MarchaV003" : Bool AT %DB90.DBX11.2, 1 s
   "ParadaV003" : Bool AT %DB90.DBX12.7, 1 s
   "BombaTorreON" : Bool AT %M69.2, 1 s
   "SirenaM5" : Bool AT %DB91.DBX0.4, 1 s
   "SirenaChillers" : Bool AT %Q68.1, 1 s
   "SirenaM6" : Bool AT %DB91.DBX0.5, 1 s
   "SirenaM7" : Bool AT %DB91.DBX0.6, 1 s
   "SirenaM8" : Bool AT %DB91.DBX0.7, 1 s
   "SirenaM9" : Bool AT %DB91.DBX1.0, 1 s
   "SirenaM10" : Bool AT %DB91.DBX1.1, 1 s
   "AlarmaNueva" : Bool AT %DB47.DBX0.0, 1 s
   "AlarmaPresente" : Bool AT %DB47.DBX0.1, 1 s
   "SinAlarmas" : Bool AT %DB47.DBX0.2, 1 s
   "AlarmaAceite-CH-ENV-CH" : Bool AT %I76.0, 1 s
   "AlarmaTemp-CH-ENV-CH" : Bool AT %I76.1, 1 s
   "RUN-CH-ENV-CH" : Bool AT %I76.2, 1 s
   "VerCh1MTA" : Bool, internal
   "VerCh2MTA" : Bool, internal
   "VerCh3MTA" : Bool, internal
   "VerCh4MTA" : Bool, internal
   "AlarmaPRUEBA" : DWord AT %DB1.DBD0, 1 s
   "Presosato" : Bool AT %I76.4, 1 s
   "CH-SOP-CH-CTC1ON" : Bool AT %I69.0, 1 s
   "CH-SOP-CH-CTC2ON" : Bool AT %I69.1, 1 s
   "CH-SOP-CH-TERM1" : Bool AT %I69.2, 1 s
   "CH-SOP-CH-TERM2" : Bool AT %I69.3, 1 s